(* CODESYS project CodeSys_main.project

Project tree, tasks and I/O mapping:
  MODULE_PLC09 : CECC-LK, Festo AG & Co. KG, order no. 574418, version 3.5.4.0
    application Application
      libraries: VisuDialogs, * (System); Solution Center Library, 3.5.8.0 (Festo Didactic SE - Customer Solution Center); CAA Real Time Clock Extern, 3.5.7.0 (CAA Technical Workgroup); CAA CiA 405, 3.5.3.0 (CAA Technical Workgroup)
      task Task (cyclic, interval t#10ms, priority 5) calls MODULE_PLC09_MAIN
      Data Types/
      Variables/
        global variables IO
        declarations NVL_PLC09_REC_FILLING
        global variables NVL_PLC09_SEND
        declarations NVL_PLC09_REC_STOPPERING
      Programs/
        program MODULE_PLC09_MAIN [ST]
      Symbols
    CANbus : CANbus, 3S - Smart Software Solutions GmbH, version 3.5.7.0
        settings: Baudrate = 1000
      CANopen_Manager : CANopen_Manager, 3S - Smart Software Solutions GmbH, version 3.5.7.20
          settings: Sync CycleTime in Microseconds = 10000; Enable Sync generation = TRUE; Synchronous Window Length = 8000; Enable Heartbeat generation = FALSE; Heartbeat Node ID = 1; CANopen NodeID = 1; ConfigVersion = 50659584
        BL20_GWBR_CANOPEN : BL20-GWBR-CANOPEN, TURCK, order no. 6827167, version Revision=16#00040017, FileVersion=4.23
            settings: General Options.Reset Node = FALSE; NODEIDSAVED = 2; SDO Timeout = 1000000; PDO_Autoconfig = TRUE; EXPERTSETTINGS = TRUE; SubIndex for reset node = 1; Emergency-General Parameters.Emergency COBID = 16#00000082; Settings.COBID = 16#00000202; Settings.Transmission Type = 16#00; Settings.available PDO-Parameter.Inhibit Time available = FALSE; Settings.available PDO-Parameter.Event Timer available = FALSE; Settings.Inhibit Time = 0; Settings.Event Timer = 0; Generic COBID = '$NODEID+16#0200'; Process by CANopenManager = TRUE; Settings.COBID = 16#00000302; Settings.Transmission Type = 16#00; Settings.available PDO-Parameter.Inhibit Time available = FALSE; Settings.available PDO-Parameter.Event Timer available = FALSE; Settings.Inhibit Time = 0; Settings.Event Timer = 0; Generic COBID = '$NODEID+16#0300'; Process by CANopenManager = TRUE; Settings.COBID = 16#00000182; Settings.Transmission Type = 16#01; Settings.available PDO-Parameter.Inhibit Time available = TRUE; Settings.available PDO-Parameter.Event Timer available = TRUE; Settings.Inhibit Time = 0; Settings.Event Timer = 0; Generic COBID = '$NODEID+16#0180'; Process by CANopenManager = TRUE; Settings.COBID = 16#00000282; Settings.Transmission Type = 16#00; Settings.available PDO-Parameter.Inhibit Time available = TRUE; Settings.available PDO-Parameter.Event Timer available = TRUE; Settings.Inhibit Time = 0; Settings.Event Timer = 0; Generic COBID = '$NODEID+16#0280'; Process by CANopenManager = TRUE; WriteOutput8Bit : Generic_BL20_4DO.Index = 16#6200 ... (307 more)
          Generic_BL20_4DO_1 : Generic BL20-4DO, TURCK, order no. 0, version Revision=16#00040017, FileVersion=4.23
              settings: Number of Params = 1; WriteOutput8Bit : Generic_BL20_4DO.Index = 16#6200; WriteOutput8Bit : Generic_BL20_4DO.Subindex = 16#01; WriteOutput8Bit : Generic_BL20_4DO.Startbit = 4; WriteOutput8Bit : Generic_BL20_4DO.Endbit = 7
              unmapped channels: WriteOutput8Bit : Generic_BL20_4DO
          Generic_BL20_4DI_1 : Generic BL20-4DI, TURCK, order no. 0, version Revision=16#00040017, FileVersion=4.23
              settings: Number of Params = 1; ReadInput8Bit : Generic_BL20_4DI.Index = 16#6000; ReadInput8Bit : Generic_BL20_4DI.Subindex = 16#01; ReadInput8Bit : Generic_BL20_4DI.Startbit = 4; ReadInput8Bit : Generic_BL20_4DI.Endbit = 7
              unmapped channels: ReadInput8Bit : Generic_BL20_4DI
          Generic_BL20_4AI : Generic BL20-4AI, TURCK, order no. 0, version Revision=16#00040017, FileVersion=4.23
              settings: Number of Params = 4; ReadAnalogueInput16Bit : Generic_BL20_4AI.Index = 16#6401; ReadAnalogueInput16Bit : Generic_BL20_4AI.Subindex = 16#01; ReadAnalogueInput16Bit : Generic_BL20_4AI.Startbit = 0; ReadAnalogueInput16Bit : Generic_BL20_4AI.Endbit = 15; ReadAnalogueInput16Bit : Generic_BL20_4AI.Index = 16#6401; ReadAnalogueInput16Bit : Generic_BL20_4AI.Subindex = 16#02; ReadAnalogueInput16Bit : Generic_BL20_4AI.Startbit = 0; ReadAnalogueInput16Bit : Generic_BL20_4AI.Endbit = 15; ReadAnalogueInput16Bit : Generic_BL20_4AI.Index = 16#6401; ReadAnalogueInput16Bit : Generic_BL20_4AI.Subindex = 16#03; ReadAnalogueInput16Bit : Generic_BL20_4AI.Startbit = 0; ReadAnalogueInput16Bit : Generic_BL20_4AI.Endbit = 15; ReadAnalogueInput16Bit : Generic_BL20_4AI.Index = 16#6401; ReadAnalogueInput16Bit : Generic_BL20_4AI.Subindex = 16#04; ReadAnalogueInput16Bit : Generic_BL20_4AI.Startbit = 0; ReadAnalogueInput16Bit : Generic_BL20_4AI.Endbit = 15
              unmapped channels: ReadAnalogueInput16Bit : Generic_BL20_4AI, ReadAnalogueInput16Bit : Generic_BL20_4AI, ReadAnalogueInput16Bit : Generic_BL20_4AI, ReadAnalogueInput16Bit : Generic_BL20_4AI
          Generic_BL20_4DO_2 : Generic BL20-4DO, TURCK, order no. 0, version Revision=16#00040017, FileVersion=4.23
              settings: Number of Params = 1; WriteOutput8Bit : Generic_BL20_4DO_2.Index = 16#6200; WriteOutput8Bit : Generic_BL20_4DO_2.Subindex = 16#02; WriteOutput8Bit : Generic_BL20_4DO_2.Startbit = 0; WriteOutput8Bit : Generic_BL20_4DO_2.Endbit = 3
              unmapped channels: WriteOutput8Bit : Generic_BL20_4DO_2
          Generic_BL20_4DO_3 : Generic BL20-4DO, TURCK, order no. 0, version Revision=16#00040017, FileVersion=4.23
              settings: Number of Params = 1; WriteOutput8Bit : Generic_BL20_4DO_2.Index = 16#6200; WriteOutput8Bit : Generic_BL20_4DO_2.Subindex = 16#02; WriteOutput8Bit : Generic_BL20_4DO_2.Startbit = 4; WriteOutput8Bit : Generic_BL20_4DO_2.Endbit = 7
              unmapped channels: WriteOutput8Bit : Generic_BL20_4DO_2
          Generic_BL20_4DO : Generic BL20-4DO, TURCK, order no. 0, version Revision=16#00040017, FileVersion=4.23
              settings: Number of Params = 1; WriteOutput8Bit : Generic_BL20_4DO.Index = 16#6200; WriteOutput8Bit : Generic_BL20_4DO.Subindex = 16#01; WriteOutput8Bit : Generic_BL20_4DO.Startbit = 0; WriteOutput8Bit : Generic_BL20_4DO.Endbit = 3
              unmapped channels: WriteOutput8Bit : Generic_BL20_4DO
          Generic_BL20_4DI : Generic BL20-4DI, TURCK, order no. 0, version Revision=16#00040017, FileVersion=4.23
              settings: Number of Params = 1; ReadInput8Bit : Generic_BL20_4DI.Index = 16#6000; ReadInput8Bit : Generic_BL20_4DI.Subindex = 16#01; ReadInput8Bit : Generic_BL20_4DI.Startbit = 0; ReadInput8Bit : Generic_BL20_4DI.Endbit = 3
              unmapped channels: ReadInput8Bit : Generic_BL20_4DI
          Generic_BL20_BR_PF : Generic BL20-BR/-PF, TURCK, order no. 0, version Revision=16#00040017, FileVersion=4.23
          Generic_BL20_2AO : Generic BL20-2AO, TURCK, order no. 0, version Revision=16#00040017, FileVersion=4.23
              settings: Number of Params = 2; WriteAnalogueOutput16 : Generic_BL20_2AO.Index = 16#6411; WriteAnalogueOutput16 : Generic_BL20_2AO.Subindex = 16#01; WriteAnalogueOutput16 : Generic_BL20_2AO.Startbit = 0; WriteAnalogueOutput16 : Generic_BL20_2AO.Endbit = 15; WriteAnalogueOutput16 : Generic_BL20_2AO.Index = 16#6411; WriteAnalogueOutput16 : Generic_BL20_2AO.Subindex = 16#02; WriteAnalogueOutput16 : Generic_BL20_2AO.Startbit = 0; WriteAnalogueOutput16 : Generic_BL20_2AO.Endbit = 15
              unmapped channels: WriteAnalogueOutput16 : Generic_BL20_2AO, WriteAnalogueOutput16 : Generic_BL20_2AO
        DTM425 : DTM425, ifm electronic gmbh, order no. DTM425, version Revision=16#00000000, FileVersion=8.2, File=DTM425.eds
            settings: NODEIDSAVED = 32; SDO Timeout = 1000000; PDO_Autoconfig = FALSE; EXPERTSETTINGS = FALSE; Emergency-General Parameters.Emergency COBID = 16#000000A0; Heartbeat-Producer Time = 200; PDO 16#1400.COBID = 16#00000220; Process by CANopenManager = TRUE; PDO 16#1401.COBID = 16#00000320; Process by CANopenManager = TRUE; PDO 16#1402.COBID = 16#00000420; Process by CANopenManager = TRUE; PDO 16#1403.COBID = 16#00000520; Process by CANopenManager = TRUE; PDO 16#1800.COBID = 16#000001A0; PDO 16#1800.Event Timer = 0; Process by CANopenManager = TRUE; PDO 16#1801.COBID = 16#000002A0; PDO 16#1801.Event Timer = 0; Process by CANopenManager = TRUE; PDO 16#1802.COBID = 16#000003A0; PDO 16#1802.Event Timer = 0; Process by CANopenManager = TRUE; PDO 16#1803.COBID = 16#000004A0; PDO 16#1803.Event Timer = 0; Process by CANopenManager = TRUE; Write Data (mappable): Write Trigger.Subindex = 16#00; Write Data (mappable): Data_sub1.Subindex = 16#01; Write Data (mappable): Data_sub2.Subindex = 16#02; Write Data (mappable): Data_sub3.Subindex = 16#03; Device Status.Subindex = 16#00; Read Data (mappable): Data_sub1.Subindex = 16#01; Read Data (mappable): Data_sub2.Subindex = 16#02; Read Data (mappable): Data_sub3.Subindex = 16#03; SDO List.Set COB-ID sync.Index = 16#1005; SDO List.Set COB-ID sync.Subindex = 16#00; SDO List.Set COB-ID sync.Value = 16#00000080; SDO List.Set COB-ID sync.Size = 32; SDO List.Set COB-ID sync.AbortIfError = FALSE; SDO List.Set COB-ID sync.JumpToLine = FALSE ... (387 more)
            unmapped channels: Write Data (mappable): Write Trigger, Write Data (mappable): Data_sub1, Write Data (mappable): Data_sub2, Write Data (mappable): Data_sub3, Device Status, Read Data (mappable): Data_sub1, Read Data (mappable): Data_sub2, Read Data (mappable): Data_sub3
    Onboard : CECC 14I/8O, Festo AG & Co. KG, version 3.4.5.5
        unmapped channels: Onboard Input, Onboard Output
      Digital Inputs
          unmapped channels: Onboard Input
      Digital Outputs
          unmapped channels: Onboard Output
  APP_FILLING : CECC-D, Festo AG & Co. KG, order no. 574415, version 3.5.4.0
    application Application
      libraries: Standard, * (System); Solution Center Library, 3.5.8.0 (Festo Didactic SE - Customer Solution Center)
      task Task (cyclic, interval t#20ms, priority 20) calls APP_FILLING_MAIN
      global variables IO
      program APP_FILLING_MAIN [ST]
      global variables NVL_FILLING_SEND
      declarations NVL_FILLING_REC_09
      declarations NVL_FILLING_REC_08
    Onboard : CECC 14I/8O, Festo AG & Co. KG, order no. 
      , version 3.4.5.5
        unmapped channels: Onboard Input, Onboard Output
      Digital Outputs
          unmapped channels: Onboard Output
      Digital Inputs
          unmapped channels: Onboard Input
  MODULE_PLC08 : CECC-LK, Festo AG & Co. KG, order no. 574418, version 3.5.4.0
    application Application
      libraries: VisuDialogs, * (System); Solution Center Library, 3.5.8.0 (Festo Didactic SE - Customer Solution Center); CAA Real Time Clock Extern, 3.5.7.0 (CAA Technical Workgroup); CAA CiA 405, 3.5.3.0 (CAA Technical Workgroup)
      task Task (cyclic, interval t#10ms, priority 5) calls MODULE_PLC08_MAIN
      Data Types/
      Variables/
        global variables IO
        global variables NVL_PLC08_SEND
        declarations NVL_PLC08_REC_STOPPERING
        declarations NVL_PLC08_REC_FILLING
      Programs/
        program MODULE_PLC08_MAIN [ST]
      Symbols
    Onboard : CECC 14I/8O, Festo AG & Co. KG, version 3.4.5.5
        unmapped channels: Onboard Input, Onboard Output
      Digital Inputs
          unmapped channels: Onboard Input
      Digital Outputs
          unmapped channels: Onboard Output
    CANbus : CANbus, 3S - Smart Software Solutions GmbH, version 3.5.7.0
        settings: Baudrate = 1000
      CANopen_Manager : CANopen_Manager, 3S - Smart Software Solutions GmbH, version 3.5.7.20
          settings: Sync CycleTime in Microseconds = 10000; Enable Sync generation = TRUE; Synchronous Window Length = 8000; Enable Heartbeat generation = FALSE; Heartbeat Node ID = 1; CANopen NodeID = 1; ConfigVersion = 50659584
        BL20_GWBR_CANOPEN : BL20-GWBR-CANOPEN, TURCK, order no. 6827167, version Revision=16#00040017, FileVersion=4.23
            settings: General Options.Reset Node = FALSE; NODEIDSAVED = 2; SDO Timeout = 1000000; PDO_Autoconfig = TRUE; EXPERTSETTINGS = TRUE; SubIndex for reset node = 1; Emergency-General Parameters.Emergency COBID = 16#00000082; Settings.COBID = 16#00000202; Settings.Transmission Type = 16#00; Settings.available PDO-Parameter.Inhibit Time available = FALSE; Settings.available PDO-Parameter.Event Timer available = FALSE; Settings.Inhibit Time = 0; Settings.Event Timer = 0; Generic COBID = '$NODEID+16#0200'; Process by CANopenManager = TRUE; Settings.COBID = 16#00000302; Settings.Transmission Type = 16#00; Settings.available PDO-Parameter.Inhibit Time available = FALSE; Settings.available PDO-Parameter.Event Timer available = FALSE; Settings.Inhibit Time = 0; Settings.Event Timer = 0; Generic COBID = '$NODEID+16#0300'; Process by CANopenManager = TRUE; Settings.COBID = 16#00000182; Settings.Transmission Type = 16#01; Settings.available PDO-Parameter.Inhibit Time available = TRUE; Settings.available PDO-Parameter.Event Timer available = TRUE; Settings.Inhibit Time = 0; Settings.Event Timer = 0; Generic COBID = '$NODEID+16#0180'; Process by CANopenManager = TRUE; Settings.COBID = 16#00000282; Settings.Transmission Type = 16#00; Settings.available PDO-Parameter.Inhibit Time available = TRUE; Settings.available PDO-Parameter.Event Timer available = TRUE; Settings.Inhibit Time = 0; Settings.Event Timer = 0; Generic COBID = '$NODEID+16#0280'; Process by CANopenManager = TRUE; WriteOutput8Bit : Generic_BL20_4DO.Index = 16#6200 ... (307 more)
          Generic_BL20_4DI : Generic BL20-4DI, TURCK, order no. 0, version Revision=16#00040017, FileVersion=4.23
              settings: Number of Params = 1; ReadInput8Bit : Generic_BL20_4DI.Index = 16#6000; ReadInput8Bit : Generic_BL20_4DI.Subindex = 16#01; ReadInput8Bit : Generic_BL20_4DI.Startbit = 0; ReadInput8Bit : Generic_BL20_4DI.Endbit = 3
              unmapped channels: ReadInput8Bit : Generic_BL20_4DI
          Generic_BL20_4DI_1 : Generic BL20-4DI, TURCK, order no. 0, version Revision=16#00040017, FileVersion=4.23
              settings: Number of Params = 1; ReadInput8Bit : Generic_BL20_4DI.Index = 16#6000; ReadInput8Bit : Generic_BL20_4DI.Subindex = 16#01; ReadInput8Bit : Generic_BL20_4DI.Startbit = 4; ReadInput8Bit : Generic_BL20_4DI.Endbit = 7
              unmapped channels: ReadInput8Bit : Generic_BL20_4DI
          Generic_BL20_BR_PF : Generic BL20-BR/-PF, TURCK, order no. 0, version Revision=16#00040017, FileVersion=4.23
          Generic_BL20_4DO : Generic BL20-4DO, TURCK, order no. 0, version Revision=16#00040017, FileVersion=4.23
              settings: Number of Params = 1; WriteOutput8Bit : Generic_BL20_4DO.Index = 16#6200; WriteOutput8Bit : Generic_BL20_4DO.Subindex = 16#01; WriteOutput8Bit : Generic_BL20_4DO.Startbit = 0; WriteOutput8Bit : Generic_BL20_4DO.Endbit = 3
              unmapped channels: WriteOutput8Bit : Generic_BL20_4DO
          Generic_BL20_4DO_1 : Generic BL20-4DO, TURCK, order no. 0, version Revision=16#00040017, FileVersion=4.23
              settings: Number of Params = 1; WriteOutput8Bit : Generic_BL20_4DO.Index = 16#6200; WriteOutput8Bit : Generic_BL20_4DO.Subindex = 16#01; WriteOutput8Bit : Generic_BL20_4DO.Startbit = 4; WriteOutput8Bit : Generic_BL20_4DO.Endbit = 7
              unmapped channels: WriteOutput8Bit : Generic_BL20_4DO
          Generic_BL20_4DO_2 : Generic BL20-4DO, TURCK, order no. 0, version Revision=16#00040017, FileVersion=4.23
              settings: Number of Params = 1; WriteOutput8Bit : Generic_BL20_4DO_2.Index = 16#6200; WriteOutput8Bit : Generic_BL20_4DO_2.Subindex = 16#02; WriteOutput8Bit : Generic_BL20_4DO_2.Startbit = 0; WriteOutput8Bit : Generic_BL20_4DO_2.Endbit = 3
              unmapped channels: WriteOutput8Bit : Generic_BL20_4DO_2
          Generic_BL20_4DO_3 : Generic BL20-4DO, TURCK, order no. 0, version Revision=16#00040017, FileVersion=4.23
              settings: Number of Params = 1; WriteOutput8Bit : Generic_BL20_4DO_2.Index = 16#6200; WriteOutput8Bit : Generic_BL20_4DO_2.Subindex = 16#02; WriteOutput8Bit : Generic_BL20_4DO_2.Startbit = 4; WriteOutput8Bit : Generic_BL20_4DO_2.Endbit = 7
              unmapped channels: WriteOutput8Bit : Generic_BL20_4DO_2
          Generic_BL20_4AI : Generic BL20-4AI, TURCK, order no. 0, version Revision=16#00040017, FileVersion=4.23
              settings: Number of Params = 4; ReadAnalogueInput16Bit : Generic_BL20_4AI.Index = 16#6401; ReadAnalogueInput16Bit : Generic_BL20_4AI.Subindex = 16#01; ReadAnalogueInput16Bit : Generic_BL20_4AI.Startbit = 0; ReadAnalogueInput16Bit : Generic_BL20_4AI.Endbit = 15; ReadAnalogueInput16Bit : Generic_BL20_4AI.Index = 16#6401; ReadAnalogueInput16Bit : Generic_BL20_4AI.Subindex = 16#02; ReadAnalogueInput16Bit : Generic_BL20_4AI.Startbit = 0; ReadAnalogueInput16Bit : Generic_BL20_4AI.Endbit = 15; ReadAnalogueInput16Bit : Generic_BL20_4AI.Index = 16#6401; ReadAnalogueInput16Bit : Generic_BL20_4AI.Subindex = 16#03; ReadAnalogueInput16Bit : Generic_BL20_4AI.Startbit = 0; ReadAnalogueInput16Bit : Generic_BL20_4AI.Endbit = 15; ReadAnalogueInput16Bit : Generic_BL20_4AI.Index = 16#6401; ReadAnalogueInput16Bit : Generic_BL20_4AI.Subindex = 16#04; ReadAnalogueInput16Bit : Generic_BL20_4AI.Startbit = 0; ReadAnalogueInput16Bit : Generic_BL20_4AI.Endbit = 15
              unmapped channels: ReadAnalogueInput16Bit : Generic_BL20_4AI, ReadAnalogueInput16Bit : Generic_BL20_4AI, ReadAnalogueInput16Bit : Generic_BL20_4AI, ReadAnalogueInput16Bit : Generic_BL20_4AI
          Generic_BL20_2AO : Generic BL20-2AO, TURCK, order no. 0, version Revision=16#00040017, FileVersion=4.23
              settings: Number of Params = 2; WriteAnalogueOutput16 : Generic_BL20_2AO.Index = 16#6411; WriteAnalogueOutput16 : Generic_BL20_2AO.Subindex = 16#01; WriteAnalogueOutput16 : Generic_BL20_2AO.Startbit = 0; WriteAnalogueOutput16 : Generic_BL20_2AO.Endbit = 15; WriteAnalogueOutput16 : Generic_BL20_2AO.Index = 16#6411; WriteAnalogueOutput16 : Generic_BL20_2AO.Subindex = 16#02; WriteAnalogueOutput16 : Generic_BL20_2AO.Startbit = 0; WriteAnalogueOutput16 : Generic_BL20_2AO.Endbit = 15
              unmapped channels: WriteAnalogueOutput16 : Generic_BL20_2AO, WriteAnalogueOutput16 : Generic_BL20_2AO
        DTM425 : DTM425, ifm electronic gmbh, order no. DTM425, version Revision=16#00000000, FileVersion=8.2, File=DTM425.eds
            settings: NODEIDSAVED = 32; SDO Timeout = 1000000; PDO_Autoconfig = FALSE; EXPERTSETTINGS = FALSE; Emergency-General Parameters.Emergency COBID = 16#000000A0; Heartbeat-Producer Time = 200; PDO 16#1400.COBID = 16#00000220; Process by CANopenManager = TRUE; PDO 16#1401.COBID = 16#00000320; Process by CANopenManager = TRUE; PDO 16#1402.COBID = 16#00000420; Process by CANopenManager = TRUE; PDO 16#1403.COBID = 16#00000520; Process by CANopenManager = TRUE; PDO 16#1800.COBID = 16#000001A0; PDO 16#1800.Event Timer = 0; Process by CANopenManager = TRUE; PDO 16#1801.COBID = 16#000002A0; PDO 16#1801.Event Timer = 0; Process by CANopenManager = TRUE; PDO 16#1802.COBID = 16#000003A0; PDO 16#1802.Event Timer = 0; Process by CANopenManager = TRUE; PDO 16#1803.COBID = 16#000004A0; PDO 16#1803.Event Timer = 0; Process by CANopenManager = TRUE; Write Data (mappable): Write Trigger.Subindex = 16#00; Write Data (mappable): Data_sub1.Subindex = 16#01; Write Data (mappable): Data_sub2.Subindex = 16#02; Write Data (mappable): Data_sub3.Subindex = 16#03; Device Status.Subindex = 16#00; Read Data (mappable): Data_sub1.Subindex = 16#01; Read Data (mappable): Data_sub2.Subindex = 16#02; Read Data (mappable): Data_sub3.Subindex = 16#03; SDO List.Set COB-ID sync.Index = 16#1005; SDO List.Set COB-ID sync.Subindex = 16#00; SDO List.Set COB-ID sync.Value = 16#00000080; SDO List.Set COB-ID sync.Size = 32; SDO List.Set COB-ID sync.AbortIfError = FALSE; SDO List.Set COB-ID sync.JumpToLine = FALSE ... (387 more)
            unmapped channels: Write Data (mappable): Write Trigger, Write Data (mappable): Data_sub1, Write Data (mappable): Data_sub2, Write Data (mappable): Data_sub3, Device Status, Read Data (mappable): Data_sub1, Read Data (mappable): Data_sub2, Read Data (mappable): Data_sub3
  APP_STOPPERING : CECC-LK, Festo AG & Co. KG, order no. 574418, version 3.5.4.0
    application Application
      libraries: Standard, * (System); Solution Center Library, 3.5.8.0 (Festo Didactic SE - Customer Solution Center)
      task Task (cyclic, interval t#20ms, priority 20) calls APP_STOPPERING_MAIN
      global variables IO
      program APP_STOPPERING_MAIN [ST]
      global variables NVL_STOPPERING_SEND
      declarations NVL_STOPPERING_REC_08
      declarations NVL_STOPPERING_REC_09
    Onboard : CECC 14I/8O, Festo AG & Co. KG, version 3.4.5.5
        unmapped channels: Onboard Input, Onboard Output
      Digital Inputs
          unmapped channels: Onboard Input
      Digital Outputs
          unmapped channels: Onboard Output
  libraries: Standard, * (System); Util, * (System); SysMem, 3.5.5.0 (System); VisuElemBase, 3.5.9.30 (System)
  5ce3da45-db07-42e7-a21c-a00fff4ed8f6|C:\Users\ggb\Documents\#PROJECTS\2016_06_29_Denmark\Visu\German.gif
  5ce3da45-db07-42e7-a21c-a00fff4ed8f6|C:\Users\ggb\Documents\#PROJECTS\2016_06_29_Denmark\Visu\Home_0.png
  5ce3da45-db07-42e7-a21c-a00fff4ed8f6|C:\Users\ggb\Documents\#PROJECTS\2016_06_29_Denmark\Visu\German.gif
  5ce3da45-db07-42e7-a21c-a00fff4ed8f6|C:\Users\ggb\Documents\#PROJECTS\2016_06_29_Denmark\Pictures\071-030_Modul Trocknen.jpg
  5ce3da45-db07-42e7-a21c-a00fff4ed8f6|C:\Users\ggb\Documents\#PROJECTS\2016_06_29_Denmark\Pictures\071-060_Kameraprüfen.jpg
  5ce3da45-db07-42e7-a21c-a00fff4ed8f6|C:\Users\ggb\Documents\#PROJECTS\2016_06_29_Denmark\Pictures\cpFactory_Bypass.png
  5ce3da45-db07-42e7-a21c-a00fff4ed8f6|C:\Users\ggb\Documents\#PROJECTS\2016_06_29_Denmark\Visu\Settings_0.png
  5ce3da45-db07-42e7-a21c-a00fff4ed8f6|C:\Users\ggb\Documents\#PROJECTS\2016_06_29_Denmark\Visu\Stopper.jpg
  5ce3da45-db07-42e7-a21c-a00fff4ed8f6|C:\Users\ggb\Documents\#PROJECTS\2016_06_29_Denmark\Visu\Parameters_1.png
  5ce3da45-db07-42e7-a21c-a00fff4ed8f6|C:\Users\ggb\Documents\#PROJECTS\2016_06_29_Denmark\Visu\RightArrow.png
  5ce3da45-db07-42e7-a21c-a00fff4ed8f6|C:\Users\ggb\Documents\#PROJECTS\2016_06_29_Denmark\Pictures\071-030_Modul Trocknen.jpg
  5ce3da45-db07-42e7-a21c-a00fff4ed8f6|C:\Users\ggb\Documents\#PROJECTS\2016_06_29_Denmark\Visu\Parameters_0.png
  5ce3da45-db07-42e7-a21c-a00fff4ed8f6|C:\Users\ggb\Documents\#PROJECTS\2016_06_29_Denmark\Visu\Stopper.jpg
  5ce3da45-db07-42e7-a21c-a00fff4ed8f6|C:\Users\ggb\Documents\#PROJECTS\2016_06_29_Denmark\Visu\Home_1.png
  5ce3da45-db07-42e7-a21c-a00fff4ed8f6|C:\Users\ggb\Documents\#PROJECTS\2016_06_29_Denmark\Pictures\071-060_Kameraprüfen.jpg
  5ce3da45-db07-42e7-a21c-a00fff4ed8f6|C:\Users\ggb\Documents\#PROJECTS\2016_06_29_Denmark\Visu\Settings_1.png
  5ce3da45-db07-42e7-a21c-a00fff4ed8f6|C:\Users\ggb\Documents\#PROJECTS\2016_06_29_Denmark\Pictures\cpFactory_Conveyor.png
  5ce3da45-db07-42e7-a21c-a00fff4ed8f6|C:\Users\ggb\Documents\#PROJECTS\2016_06_29_Denmark\Pictures\071-050a_Bohren EA.jpg
  5ce3da45-db07-42e7-a21c-a00fff4ed8f6|C:\Users\ggb\Documents\#PROJECTS\2016_06_29_Denmark\Visu\Manual_1.png
  5ce3da45-db07-42e7-a21c-a00fff4ed8f6|C:\Users\ggb\Documents\#PROJECTS\2016_06_29_Denmark\Pictures\071-060_Kameraprüfen.jpg
  5ce3da45-db07-42e7-a21c-a00fff4ed8f6|C:\Users\ggb\Documents\#PROJECTS\2016_06_29_Denmark\Visu\Settings_1.png
  5ce3da45-db07-42e7-a21c-a00fff4ed8f6|C:\Users\ggb\Documents\#PROJECTS\2016_06_29_Denmark\Visu\RightArrow.png
  5ce3da45-db07-42e7-a21c-a00fff4ed8f6|C:\Users\ggb\Documents\#PROJECTS\2016_06_29_Denmark\Visu\Manual_0.png
  5ce3da45-db07-42e7-a21c-a00fff4ed8f6|C:\Users\ggb\Documents\#PROJECTS\2016_06_29_Denmark\Pictures\071-030_Modul Trocknen.jpg
  5ce3da45-db07-42e7-a21c-a00fff4ed8f6|C:\Users\ggb\Documents\#PROJECTS\2016_06_29_Denmark\Visu\German.gif
  5ce3da45-db07-42e7-a21c-a00fff4ed8f6|C:\Users\ggb\Documents\#PROJECTS\2016_06_29_Denmark\Visu\Stopper.jpg
  5ce3da45-db07-42e7-a21c-a00fff4ed8f6|C:\Users\ggb\Documents\#PROJECTS\2016_06_29_Denmark\Visu\RightArrow_Bold.png
  5ce3da45-db07-42e7-a21c-a00fff4ed8f6|C:\Users\ggb\Documents\#PROJECTS\2016_06_29_Denmark\Visu\FESTO.png
  5ce3da45-db07-42e7-a21c-a00fff4ed8f6|C:\Users\ggb\Documents\#PROJECTS\2016_06_29_Denmark\Visu\Stopper.jpg
  5ce3da45-db07-42e7-a21c-a00fff4ed8f6|C:\Users\ggb\Documents\#PROJECTS\2016_06_29_Denmark\Visu\Parameters_1.png
  5ce3da45-db07-42e7-a21c-a00fff4ed8f6|C:\Users\ggb\Documents\#PROJECTS\2016_06_29_Denmark\Visu\Parameters_0.png
  5ce3da45-db07-42e7-a21c-a00fff4ed8f6|C:\Users\ggb\Documents\#PROJECTS\2016_06_29_Denmark\Pictures\cpFactory_Bypass.png
  5ce3da45-db07-42e7-a21c-a00fff4ed8f6|C:\Users\ggb\Documents\#PROJECTS\2016_06_29_Denmark\Pictures\071-030_Modul Trocknen.jpg
  5ce3da45-db07-42e7-a21c-a00fff4ed8f6|C:\Users\ggb\Documents\#PROJECTS\2016_06_29_Denmark\Visu\CheckBox_1.png
  5ce3da45-db07-42e7-a21c-a00fff4ed8f6|C:\Users\ggb\Documents\#PROJECTS\2016_06_29_Denmark\Visu\Settings_0.png
  5ce3da45-db07-42e7-a21c-a00fff4ed8f6|C:\Users\ggb\Documents\#PROJECTS\2016_06_29_Denmark\Visu\Plus.png
  5ce3da45-db07-42e7-a21c-a00fff4ed8f6|C:\Users\ggb\Documents\#PROJECTS\2016_06_29_Denmark\Visu\CheckBox_0.png
  5ce3da45-db07-42e7-a21c-a00fff4ed8f6|C:\Users\ggb\Documents\#PROJECTS\2016_06_29_Denmark\Visu\Manual_0.png
  5ce3da45-db07-42e7-a21c-a00fff4ed8f6|C:\Users\ggb\Documents\#PROJECTS\2016_06_29_Denmark\Visu\Manual_1.png
  5ce3da45-db07-42e7-a21c-a00fff4ed8f6|C:\Users\ggb\Documents\#PROJECTS\2016_06_29_Denmark\Visu\Stopper.jpg
  5ce3da45-db07-42e7-a21c-a00fff4ed8f6|C:\Users\ggb\Documents\#PROJECTS\2016_06_29_Denmark\Visu\Settings_1.png
  5ce3da45-db07-42e7-a21c-a00fff4ed8f6|C:\Users\ggb\Documents\#PROJECTS\2016_06_29_Denmark\Visu\Manual_1.png
  5ce3da45-db07-42e7-a21c-a00fff4ed8f6|C:\Users\ggb\Documents\#PROJECTS\2016_06_29_Denmark\Visu\RightArrow.png
  5ce3da45-db07-42e7-a21c-a00fff4ed8f6|C:\Users\ggb\Documents\#PROJECTS\2016_06_29_Denmark\Pictures\cpFactory_Bypass.png
  5ce3da45-db07-42e7-a21c-a00fff4ed8f6|C:\Users\ggb\Documents\#PROJECTS\2016_06_29_Denmark\Visu\Home_0.png
  5ce3da45-db07-42e7-a21c-a00fff4ed8f6|C:\Users\ggb\Documents\#PROJECTS\2016_06_29_Denmark\Pictures\071-060_Kameraprüfen.jpg
  5ce3da45-db07-42e7-a21c-a00fff4ed8f6|C:\Users\ggb\Documents\#PROJECTS\2016_06_29_Denmark\Pictures\071-050a_Bohren EA.jpg
  5ce3da45-db07-42e7-a21c-a00fff4ed8f6|C:\Users\ggb\Documents\#PROJECTS\2016_06_29_Denmark\Visu\Settings_1.png
  5ce3da45-db07-42e7-a21c-a00fff4ed8f6|C:\Users\ggb\Documents\#PROJECTS\2016_06_29_Denmark\Visu\RightArrow.png
  5ce3da45-db07-42e7-a21c-a00fff4ed8f6|C:\Users\ggb\Documents\#PROJECTS\2016_06_29_Denmark\Visu\Home_1.png
  5ce3da45-db07-42e7-a21c-a00fff4ed8f6|C:\Users\ggb\Documents\#PROJECTS\2016_06_29_Denmark\Visu\English.gif
  5ce3da45-db07-42e7-a21c-a00fff4ed8f6|C:\Users\ggb\Documents\#PROJECTS\2016_06_29_Denmark\Visu\LeftArrow_Bold.png
  5ce3da45-db07-42e7-a21c-a00fff4ed8f6|C:\Users\ggb\Documents\#PROJECTS\2016_06_29_Denmark\Visu\Plus.png
  5ce3da45-db07-42e7-a21c-a00fff4ed8f6|C:\Users\ggb\Documents\#PROJECTS\2016_06_29_Denmark\Pictures\071-050a_Bohren EA.jpg
  5ce3da45-db07-42e7-a21c-a00fff4ed8f6|C:\Users\ggb\Documents\#PROJECTS\2016_06_29_Denmark\Visu\RightArrow.png
  5ce3da45-db07-42e7-a21c-a00fff4ed8f6|C:\Users\ggb\Documents\#PROJECTS\2016_06_29_Denmark\Visu\Manual_1.png
  5ce3da45-db07-42e7-a21c-a00fff4ed8f6|C:\Users\ggb\Documents\#PROJECTS\2016_06_29_Denmark\Visu\German.gif
  5ce3da45-db07-42e7-a21c-a00fff4ed8f6|C:\Users\ggb\Documents\#PROJECTS\2016_06_29_Denmark\Visu\CheckBox_1.png
  5ce3da45-db07-42e7-a21c-a00fff4ed8f6|C:\Users\ggb\Documents\#PROJECTS\2016_06_29_Denmark\Pictures\071-050a_Bohren EA.jpg
  5ce3da45-db07-42e7-a21c-a00fff4ed8f6|C:\Users\ggb\Documents\#PROJECTS\2016_06_29_Denmark\Visu\LeftArrow_Bold.png
  5ce3da45-db07-42e7-a21c-a00fff4ed8f6|C:\Users\ggb\Documents\#PROJECTS\2016_06_29_Denmark\Visu\Parameters_0.png
  5ce3da45-db07-42e7-a21c-a00fff4ed8f6|C:\Users\ggb\Documents\#PROJECTS\2016_06_29_Denmark\Visu\Home_0.png
  5ce3da45-db07-42e7-a21c-a00fff4ed8f6|C:\Users\ggb\Documents\#PROJECTS\2016_06_29_Denmark\Visu\Settings_0.png
  5ce3da45-db07-42e7-a21c-a00fff4ed8f6|C:\Users\ggb\Documents\#PROJECTS\2016_06_29_Denmark\Visu\Settings_1.png
  5ce3da45-db07-42e7-a21c-a00fff4ed8f6|C:\Users\ggb\Documents\#PROJECTS\2016_06_29_Denmark\Pictures\cpFactory_Conveyor.png
  5ce3da45-db07-42e7-a21c-a00fff4ed8f6|C:\Users\ggb\Documents\#PROJECTS\2016_06_29_Denmark\Pictures\071-046b_Magazin.jpg
  5ce3da45-db07-42e7-a21c-a00fff4ed8f6|C:\Users\ggb\Documents\#PROJECTS\2016_06_29_Denmark\Visu\Home_0.png
  5ce3da45-db07-42e7-a21c-a00fff4ed8f6|C:\Users\ggb\Documents\#PROJECTS\2016_06_29_Denmark\Visu\English.gif
  5ce3da45-db07-42e7-a21c-a00fff4ed8f6|C:\Users\ggb\Documents\#PROJECTS\2016_06_29_Denmark\Visu\Manual_0.png
  5ce3da45-db07-42e7-a21c-a00fff4ed8f6|C:\Users\ggb\Documents\#PROJECTS\2016_06_29_Denmark\Visu\Parameters_0.png
  5ce3da45-db07-42e7-a21c-a00fff4ed8f6|C:\Users\ggb\Documents\#PROJECTS\2016_06_29_Denmark\Visu\CheckBox_0.png
  5ce3da45-db07-42e7-a21c-a00fff4ed8f6|C:\Users\ggb\Documents\#PROJECTS\2016_06_29_Denmark\Visu\Settings_0.png
  5ce3da45-db07-42e7-a21c-a00fff4ed8f6|C:\Users\ggb\Documents\#PROJECTS\2016_06_29_Denmark\Pictures\cpFactory_Bypass.png
  5ce3da45-db07-42e7-a21c-a00fff4ed8f6|C:\Users\ggb\Documents\#PROJECTS\2016_06_29_Denmark\Visu\CheckBox_0.png
  5ce3da45-db07-42e7-a21c-a00fff4ed8f6|C:\Users\ggb\Documents\#PROJECTS\2016_06_29_Denmark\Visu\Parameters_0.png
  5ce3da45-db07-42e7-a21c-a00fff4ed8f6|C:\Users\ggb\Documents\#PROJECTS\2016_06_29_Denmark\Pictures\071-050a_Bohren EA.jpg
  5ce3da45-db07-42e7-a21c-a00fff4ed8f6|C:\Users\ggb\Documents\#PROJECTS\2016_06_29_Denmark\Visu\Parameters_1.png
  5ce3da45-db07-42e7-a21c-a00fff4ed8f6|C:\Users\ggb\Documents\#PROJECTS\2016_06_29_Denmark\Visu\Manual_0.png
  5ce3da45-db07-42e7-a21c-a00fff4ed8f6|C:\Users\ggb\Documents\#PROJECTS\2016_06_29_Denmark\Pictures\071-030_Modul Trocknen.jpg
  5ce3da45-db07-42e7-a21c-a00fff4ed8f6|C:\Users\ggb\Documents\#PROJECTS\2016_06_29_Denmark\Pictures\071-050a_Bohren EA.jpg
  5ce3da45-db07-42e7-a21c-a00fff4ed8f6|C:\Users\ggb\Documents\#PROJECTS\2016_06_29_Denmark\Pictures\cpFactory_Conveyor.png
  5ce3da45-db07-42e7-a21c-a00fff4ed8f6|C:\Users\ggb\Documents\#PROJECTS\2016_06_29_Denmark\Visu\RightArrow.png
  5ce3da45-db07-42e7-a21c-a00fff4ed8f6|C:\Users\ggb\Documents\#PROJECTS\2016_06_29_Denmark\Visu\Plus.png
  5ce3da45-db07-42e7-a21c-a00fff4ed8f6|C:\Users\ggb\Documents\#PROJECTS\2016_06_29_Denmark\Visu\Manual_0.png
  5ce3da45-db07-42e7-a21c-a00fff4ed8f6|C:\Users\ggb\Documents\#PROJECTS\2016_06_29_Denmark\Visu\Home_1.png
  5ce3da45-db07-42e7-a21c-a00fff4ed8f6|C:\Users\ggb\Documents\#PROJECTS\2016_06_29_Denmark\Visu\RightArrow.png
  5ce3da45-db07-42e7-a21c-a00fff4ed8f6|C:\Users\ggb\Documents\#PROJECTS\2016_06_29_Denmark\Visu\Settings_0.png
  5ce3da45-db07-42e7-a21c-a00fff4ed8f6|C:\Users\ggb\Documents\#PROJECTS\2016_06_29_Denmark\Visu\Plus.png
  5ce3da45-db07-42e7-a21c-a00fff4ed8f6|C:\Users\ggb\Documents\#PROJECTS\2016_06_29_Denmark\Pictures\cpFactory_Conveyor.png
  5ce3da45-db07-42e7-a21c-a00fff4ed8f6|C:\Users\ggb\Documents\#PROJECTS\2016_06_29_Denmark\Visu\English.gif
  5ce3da45-db07-42e7-a21c-a00fff4ed8f6|C:\Users\ggb\Documents\#PROJECTS\2016_06_29_Denmark\Pictures\071-060_Kameraprüfen.jpg
  5ce3da45-db07-42e7-a21c-a00fff4ed8f6|C:\Users\ggb\Documents\#PROJECTS\2016_06_29_Denmark\Visu\RightArrow.png
  5ce3da45-db07-42e7-a21c-a00fff4ed8f6|C:\Users\ggb\Documents\#PROJECTS\2016_06_29_Denmark\Pictures\071-046b_Magazin.jpg
  5ce3da45-db07-42e7-a21c-a00fff4ed8f6|C:\Users\ggb\Documents\#PROJECTS\2016_06_29_Denmark\Pictures\071-030_Modul Trocknen.jpg
  5ce3da45-db07-42e7-a21c-a00fff4ed8f6|C:\Users\ggb\Documents\#PROJECTS\2016_06_29_Denmark\Visu\Home_0.png
  5ce3da45-db07-42e7-a21c-a00fff4ed8f6|C:\Users\ggb\Documents\#PROJECTS\2016_06_29_Denmark\Pictures\071-060_Kameraprüfen.jpg
  5ce3da45-db07-42e7-a21c-a00fff4ed8f6|C:\Users\ggb\Documents\#PROJECTS\2016_06_29_Denmark\Visu\Manual_1.png
  5ce3da45-db07-42e7-a21c-a00fff4ed8f6|C:\Users\ggb\Documents\#PROJECTS\2016_06_29_Denmark\Visu\Manual_0.png
  5ce3da45-db07-42e7-a21c-a00fff4ed8f6|C:\Users\ggb\Documents\#PROJECTS\2016_06_29_Denmark\Visu\FESTO.png
  5ce3da45-db07-42e7-a21c-a00fff4ed8f6|C:\Users\ggb\Documents\#PROJECTS\2016_06_29_Denmark\Visu\Parameters_1.png
  5ce3da45-db07-42e7-a21c-a00fff4ed8f6|C:\Users\ggb\Documents\#PROJECTS\2016_06_29_Denmark\Visu\Plus.png
  5ce3da45-db07-42e7-a21c-a00fff4ed8f6|C:\Users\ggb\Documents\#PROJECTS\2016_06_29_Denmark\Pictures\cpFactory_Bypass.png
  5ce3da45-db07-42e7-a21c-a00fff4ed8f6|C:\Users\ggb\Documents\#PROJECTS\2016_06_29_Denmark\Pictures\071-050a_Bohren EA.jpg
  5ce3da45-db07-42e7-a21c-a00fff4ed8f6|C:\Users\ggb\Documents\#PROJECTS\2016_06_29_Denmark\Visu\FESTO.png
  5ce3da45-db07-42e7-a21c-a00fff4ed8f6|C:\Users\ggb\Documents\#PROJECTS\2016_06_29_Denmark\Visu\Home_1.png
  5ce3da45-db07-42e7-a21c-a00fff4ed8f6|C:\Users\ggb\Documents\#PROJECTS\2016_06_29_Denmark\Visu\Parameters_0.png
  5ce3da45-db07-42e7-a21c-a00fff4ed8f6|C:\Users\ggb\Documents\#PROJECTS\2016_06_29_Denmark\Visu\Parameters_1.png
  5ce3da45-db07-42e7-a21c-a00fff4ed8f6|C:\Users\ggb\Documents\#PROJECTS\2016_06_29_Denmark\Pictures\cpFactory_Bypass.png